VERSION : 0.1
   VAR_INPUT
      Ir_Pos_1 : Bool;   // Comando Mover Cilindro a Posición 1, activar constantemente
      Ir_Pos_2 : Bool;   // Comando Mover Cilindro a Posición 2, activar constantemente
      Conf_Pos_1 : Bool;   // Confirmación Cilindro en Posición 1
      Conf_Pos_2 : Bool;   // Confirmación Cilindro en Posición 2
      T_Conf : Time := T#10s;   // Tiempo admisible para confirmación de posición
      T_ON : Time;   // Duración accionamiento salida [0 = constantemente]
   END_VAR
   VAR_OUTPUT
      Pos_1 : Bool;   // Orden Mover Cilindro a Posición 1
      Pos_2 : Bool;   // Orden Mover Cilindro a Posición 2
      ERROR : Int;   // 0 = Sin Error, 1 = Error Programación, 2 = Error Doble Confirmación, 3 = Error Confirmación Pos_1, 4 = Error Confirmación Pos_2, 5 = Sin Confirmaciones
   END_VAR
   VAR
      IEC_Timer_0_Instance : IEC_TIMER;
      IEC_Timer_0_Instance_1 : IEC_TIMER;
      IEC_Timer_0_Instance_2 : IEC_TIMER;
      IEC_Timer_0_Instance_3 : IEC_TIMER;
      IEC_Timer_0_Instance_4 : IEC_TIMER;
   END_VAR
   VAR_TEMP
      Aux_1 : Bool;   // Auxiliar 1
      Aux_2 : Bool;   // Auxiliar 2
      Aux_ERROR : Int;   // Auxiliar ERROR
   END_VAR
BEGIN

REGION Network 1: Auxiliar 1
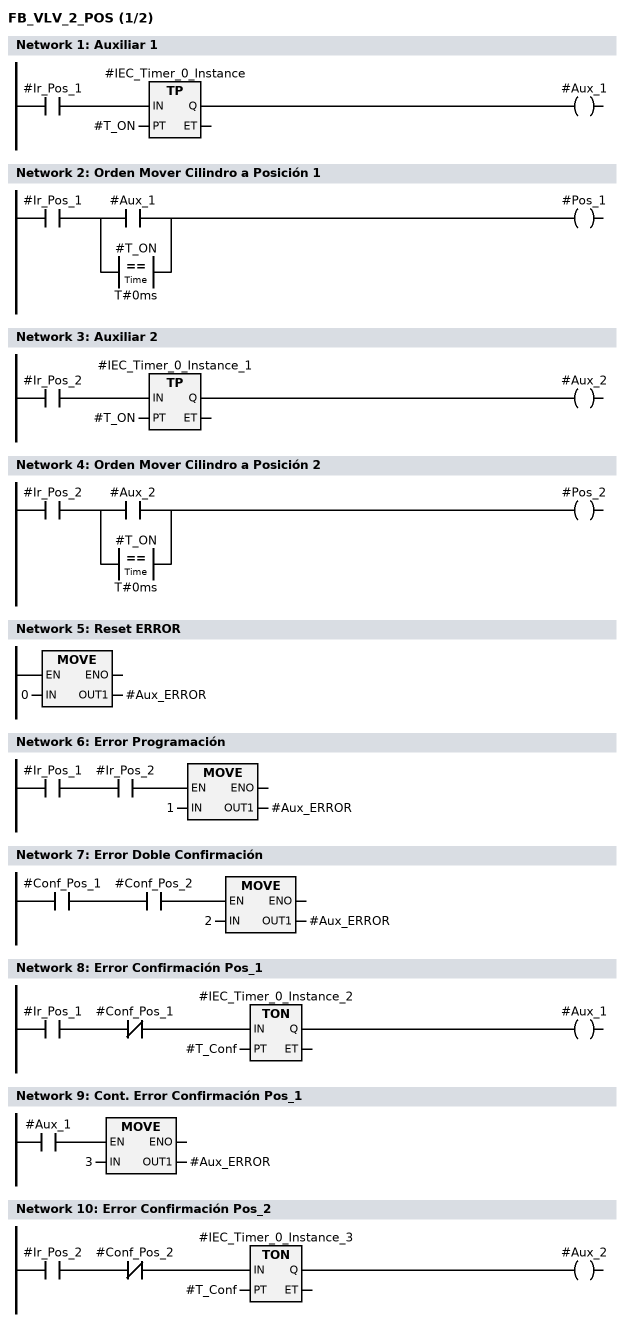
   #IEC_Timer_0_Instance.TP(IN := #Ir_Pos_1, PT := #T_ON);
   #Aux_1 := #IEC_Timer_0_Instance.Q;
END_REGION

REGION Network 2: Orden Mover Cilindro a Posición 1
   RUNG wire#powerrail
      Contact( #Ir_Pos_1 )
      wire#w1
      Contact( #Aux_1 )
      wire#w2
      Coil( #Pos_1 )
   END_RUNG
   RUNG wire#w1
      { S7_Templates := "SrcType := Time" } EQ_Contact(in1 := #T_ON, in2 := T#0ms)
   END_RUNG wire#w2
   // the same network as SCL:
   #Pos_1 := #Ir_Pos_1 AND (#Aux_1 OR (#T_ON = T#0ms));
END_REGION

REGION Network 3: Auxiliar 2
   #IEC_Timer_0_Instance_1.TP(IN := #Ir_Pos_2, PT := #T_ON);
   #Aux_2 := #IEC_Timer_0_Instance_1.Q;
END_REGION

REGION Network 4: Orden Mover Cilindro a Posición 2
   RUNG wire#powerrail
      Contact( #Ir_Pos_2 )
      wire#w1
      Contact( #Aux_2 )
      wire#w2
      Coil( #Pos_2 )
   END_RUNG
   RUNG wire#w1
      { S7_Templates := "SrcType := Time" } EQ_Contact(in1 := #T_ON, in2 := T#0ms)
   END_RUNG wire#w2
   // the same network as SCL:
   #Pos_2 := #Ir_Pos_2 AND (#Aux_2 OR (#T_ON = T#0ms));
END_REGION

REGION Network 5: Reset ERROR
   RUNG wire#powerrail
      { S7_GenerateENO := "TRUE" } Move(in := 0, out1 => #Aux_ERROR)
   END_RUNG
   // the same network as SCL:
   #Aux_ERROR := 0;
END_REGION

REGION Network 6: Error Programación
   RUNG wire#powerrail
      Contact( #Ir_Pos_1 )
      Contact( #Ir_Pos_2 )
      { S7_GenerateENO := "TRUE" } Move(in := 1, out1 => #Aux_ERROR)
   END_RUNG
   // the same network as SCL:
   IF #Ir_Pos_1 AND #Ir_Pos_2 THEN #Aux_ERROR := 1; END_IF;
END_REGION

REGION Network 7: Error Doble Confirmación
   RUNG wire#powerrail
      Contact( #Conf_Pos_1 )
      Contact( #Conf_Pos_2 )
      { S7_GenerateENO := "TRUE" } Move(in := 2, out1 => #Aux_ERROR)
   END_RUNG
   // the same network as SCL:
   IF #Conf_Pos_1 AND #Conf_Pos_2 THEN #Aux_ERROR := 2; END_IF;
END_REGION

REGION Network 8: Error Confirmación Pos_1
   #IEC_Timer_0_Instance_2.TON(IN := #Ir_Pos_1 AND NOT #Conf_Pos_1, PT := #T_Conf);
   #Aux_1 := #IEC_Timer_0_Instance_2.Q;
END_REGION

REGION Network 9: Cont. Error Confirmación Pos_1
   RUNG wire#powerrail
      Contact( #Aux_1 )
      { S7_GenerateENO := "TRUE" } Move(in := 3, out1 => #Aux_ERROR)
   END_RUNG
   // the same network as SCL:
   IF #Aux_1 THEN #Aux_ERROR := 3; END_IF;
END_REGION

REGION Network 10: Error Confirmación Pos_2
   #IEC_Timer_0_Instance_3.TON(IN := #Ir_Pos_2 AND NOT #Conf_Pos_2, PT := #T_Conf);
   #Aux_2 := #IEC_Timer_0_Instance_3.Q;
END_REGION

REGION Network 11: Cont. Error Confirmación Pos_2
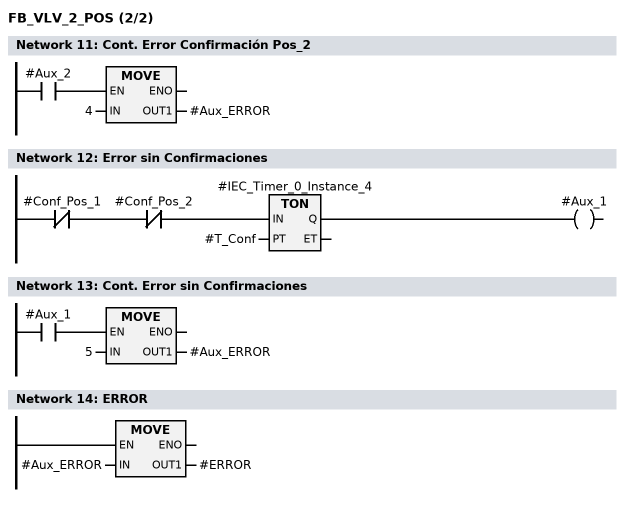
   RUNG wire#powerrail
      Contact( #Aux_2 )
      { S7_GenerateENO := "TRUE" } Move(in := 4, out1 => #Aux_ERROR)
   END_RUNG
   // the same network as SCL:
   IF #Aux_2 THEN #Aux_ERROR := 4; END_IF;
END_REGION

REGION Network 12: Error sin Confirmaciones
   #IEC_Timer_0_Instance_4.TON(IN := NOT #Conf_Pos_1 AND NOT #Conf_Pos_2, PT := #T_Conf);
   #Aux_1 := #IEC_Timer_0_Instance_4.Q;
END_REGION

REGION Network 13: Cont. Error sin Confirmaciones
   RUNG wire#powerrail
      Contact( #Aux_1 )
      { S7_GenerateENO := "TRUE" } Move(in := 5, out1 => #Aux_ERROR)
   END_RUNG
   // the same network as SCL:
   IF #Aux_1 THEN #Aux_ERROR := 5; END_IF;
END_REGION

REGION Network 14: ERROR
   RUNG wire#powerrail
      { S7_GenerateENO := "TRUE" } Move(in := #Aux_ERROR, out1 => #ERROR)
   END_RUNG
   // the same network as SCL:
   #ERROR := #Aux_ERROR;
END_REGION
END_FUNCTION_BLOCK

FUNCTION "MAQ_EST_32" : Void   // FC7, SCL
TITLE = Máquina de Estados 32
{ S7_Optimized_Access := 'TRUE' }
AUTHOR : FRD
FAMILY : MTA
NAME : MaqEst32
VERSION : 1.0
// KNOW_HOW_PROTECT  Máquina de estados de hasta 32 estados.
   VAR_INPUT
      Concatenadoras : DWord;   // Próximo estado de transición normal
      Prioritarias : DWord;   // Próximo estado de transición forzada
   END_VAR
   VAR_OUTPUT
      Error_Concatenadoras : Bool;   // Error en la programación de las Concatenadoras
      Error_Prioritarias : Bool;   // Error en la programación de las Prioritarias
   END_VAR
   VAR_IN_OUT
      Estado : DWord;   // Estado actual
   END_VAR
   VAR_TEMP
      Concat_Int : Int;   // Auxiliar INT para verificar las Concatenadoras
      Priorit_Int : Int;   // Auxiliar INT para verificar las Prioritarias
      Concat_Dword : DWord;   // Auxiliar DWORD para verificar las Concatenadoras
      Priorit_Dword : DWord;   // Auxiliar DWORD para verificar las Prioritarias
      Activar_Concat : Bool;   // Bit que indica Concatenadoras correctas
      Activar_Priorit : Bool;   // Bit que indica Prioritarias correctas
      Falla_Concat : Bool;   // Bit que indica falla en Concatenadoras
      Falla_Priorit : Bool;   // Bit que indica falla en Prioritarias
   END_VAR
BEGIN
   #Falla_Concat := 0;
   #Activar_Concat := 0;
   #Falla_Priorit := 0;
   #Activar_Priorit := 0; 
   #Error_Concatenadoras := 0;
   #Error_Prioritarias := 0;

   IF #Concatenadoras <> 0 THEN     //Evaluar Concatenadoras si son distintas de "0"

    #Concat_Int := ENCO(IN := #Concatenadoras );  //Convierte posición_DWORD en INT (0 a 31), lee el LSb

    #Concat_Dword := DECO(IN := INT_TO_UINT(#Concat_Int));//Convierte INT en posición_DWORD (1 a 32)

    IF #Concatenadoras = #Concat_Dword THEN  //Si son iguales, había sólo un bit en "1"

     #Activar_Concat := 1;    //Concatenadora correcta

    ELSE

     #Falla_Concat := 1;    //Falla en Concatenadora

    END_IF;

   END_IF;

   IF #Prioritarias <> 0 THEN     //Evaluar Prioritarias si son distintas de "0"

    #Priorit_Int := ENCO(IN := #Prioritarias);  //Convierte posición_DWORD en INT (0 a 31), lee el LSb

    #Priorit_Dword := DECO(IN := INT_TO_UINT(#Priorit_Int));//Convierte INT en posición_DWORD (1 a 32)

    IF #Prioritarias = #Priorit_Dword THEN  //Si son iguales, había sólo un bit en "1"

     #Activar_Priorit := 1;   //Prioritaria correcta

    ELSE

     #Falla_Priorit := 1;    //Falla en Prioritaria

    END_IF;

   END_IF;

   IF NOT(#Falla_Priorit OR #Falla_Concat) THEN  //Si no hay falla de Prioritaria ni de Concatenadora

    IF #Activar_Priorit THEN    //Si hay que asignar Prioritarias

     #Estado := #Prioritarias;

    ELSE

     IF #Activar_Concat THEN   //Si hay que asignar Concatenadoras

      #Estado := #Concatenadoras;

     END_IF;

    END_IF;

   ELSE

    IF #Falla_Concat THEN     //Si hay falla de Concatenadoras

     #Error_Concatenadoras := 1;    //Activar Error_Concatenadoras

    END_IF;

    IF #Falla_Priorit THEN    //Si hay falla de Prioritarias

     #Error_Prioritarias := 1;    //Activar Error_Prioritarias

    END_IF;

   END_IF;
END_FUNCTION

// folder: INCIDENTES

FUNCTION_BLOCK "FB_INC_GENERAL"   // FB500, LAD
TITLE = ALARMAS GENERAL
{ S7_Optimized_Access := 'FALSE' }
VERSION : 0.1
   VAR
      Alarma_On : Bool;
   END_VAR
BEGIN

REGION Network 1: Alarma 0 - Protecciones abiertas
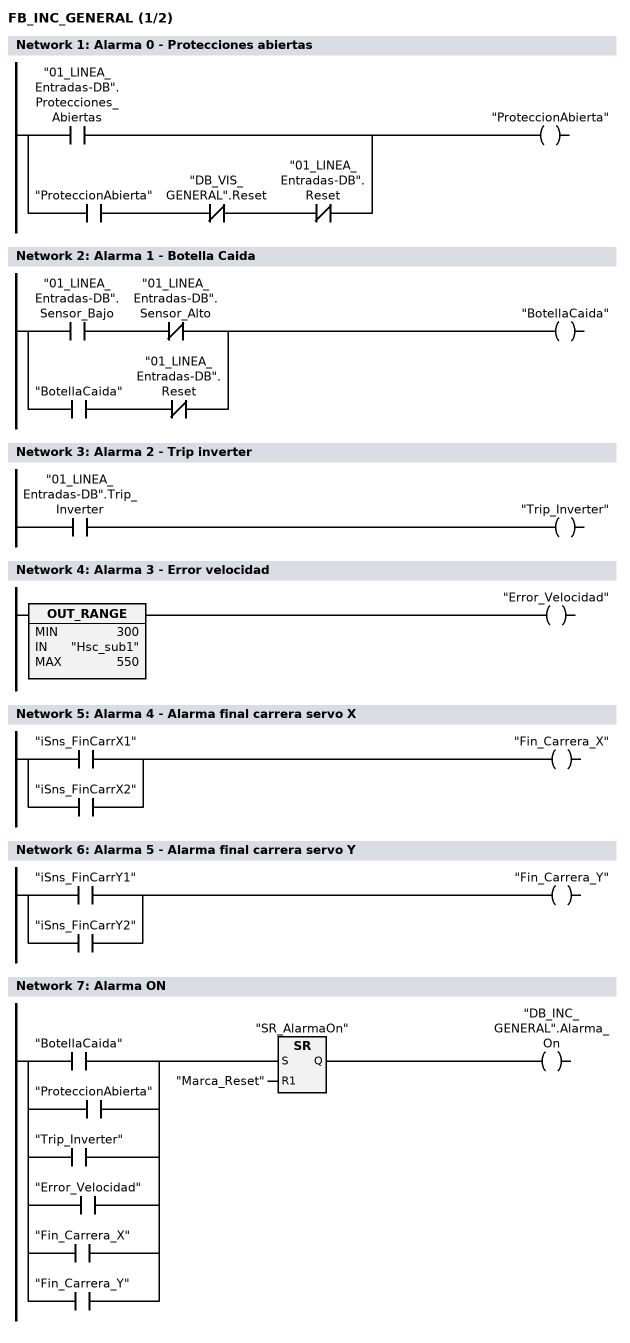
   RUNG wire#powerrail
      Contact( "01_LINEA_Entradas-DB".Protecciones_Abiertas )
      wire#w1
      Coil( "ProteccionAbierta" )
   END_RUNG
   RUNG wire#powerrail
      Contact( "ProteccionAbierta" )
      I_Contact( "DB_VIS_GENERAL".Reset )
      I_Contact( "01_LINEA_Entradas-DB".Reset )
   END_RUNG wire#w1
   // the same network as SCL:
   "ProteccionAbierta" := "01_LINEA_Entradas-DB".Protecciones_Abiertas OR ("ProteccionAbierta" AND NOT "DB_VIS_GENERAL".Reset AND NOT "01_LINEA_Entradas-DB".Reset);
END_REGION

REGION Network 2: Alarma 1 - Botella Caida
   RUNG wire#powerrail
      Contact( "01_LINEA_Entradas-DB".Sensor_Bajo )
      I_Contact( "01_LINEA_Entradas-DB".Sensor_Alto )
      wire#w1
      Coil( "BotellaCaida" )
   END_RUNG
   RUNG wire#powerrail
      Contact( "BotellaCaida" )
      I_Contact( "01_LINEA_Entradas-DB".Reset )
   END_RUNG wire#w1
   // the same network as SCL:
   "BotellaCaida" := ("01_LINEA_Entradas-DB".Sensor_Bajo AND NOT "01_LINEA_Entradas-DB".Sensor_Alto) OR ("BotellaCaida" AND NOT "01_LINEA_Entradas-DB".Reset);
END_REGION

REGION Network 3: Alarma 2 - Trip inverter
   RUNG wire#powerrail
      Contact( "01_LINEA_Entradas-DB".Trip_Inverter )
      Coil( "Trip_Inverter" )
   END_RUNG
   // the same network as SCL:
   "Trip_Inverter" := "01_LINEA_Entradas-DB".Trip_Inverter;
END_REGION

REGION Network 4: Alarma 3 - Error velocidad
   "Error_Velocidad" := ("Hsc_sub1" < 300) OR ("Hsc_sub1" > 550);
END_REGION

REGION Network 5: Alarma 4 - Alarma final carrera servo X
   RUNG wire#powerrail
      Contact( "iSns_FinCarrX1" )
      wire#w1
      Coil( "Fin_Carrera_X" )
   END_RUNG
   RUNG wire#powerrail
      Contact( "iSns_FinCarrX2" )
   END_RUNG wire#w1
   // the same network as SCL:
   "Fin_Carrera_X" := "iSns_FinCarrX1" OR "iSns_FinCarrX2";
END_REGION

REGION Network 6: Alarma 5 - Alarma final carrera servo Y
   RUNG wire#powerrail
      Contact( "iSns_FinCarrY1" )
      wire#w1
      Coil( "Fin_Carrera_Y" )
   END_RUNG
   RUNG wire#powerrail
      Contact( "iSns_FinCarrY2" )
   END_RUNG wire#w1
   // the same network as SCL:
   "Fin_Carrera_Y" := "iSns_FinCarrY1" OR "iSns_FinCarrY2";
END_REGION

REGION Network 7: Alarma ON
   RUNG wire#powerrail
      Contact( "BotellaCaida" )
      wire#w1
      S_SR(operand := "SR_AlarmaOn", r1 := "Marca_Reset")
      Coil( "DB_INC_GENERAL".Alarma_On )
   END_RUNG
   RUNG wire#powerrail
      Contact( "ProteccionAbierta" )
   END_RUNG wire#w1
   RUNG wire#powerrail
      Contact( "Trip_Inverter" )
   END_RUNG wire#w1
   RUNG wire#powerrail
      Contact( "Error_Velocidad" )
   END_RUNG wire#w1
   RUNG wire#powerrail
      Contact( "Fin_Carrera_X" )
   END_RUNG wire#w1
   RUNG wire#powerrail
      Contact( "Fin_Carrera_Y" )
   END_RUNG wire#w1
   // the same network as SCL:
   IF "BotellaCaida" OR "ProteccionAbierta" OR "Trip_Inverter" OR "Error_Velocidad" OR "Fin_Carrera_X" OR "Fin_Carrera_Y" THEN
       "SR_AlarmaOn" := TRUE;   // SR flip-flop
   END_IF;
   IF "Marca_Reset" THEN "SR_AlarmaOn" := FALSE; END_IF;
   "DB_INC_GENERAL".Alarma_On := "SR_AlarmaOn";
END_REGION

REGION Network 8: Encendido Semaforo Rojo
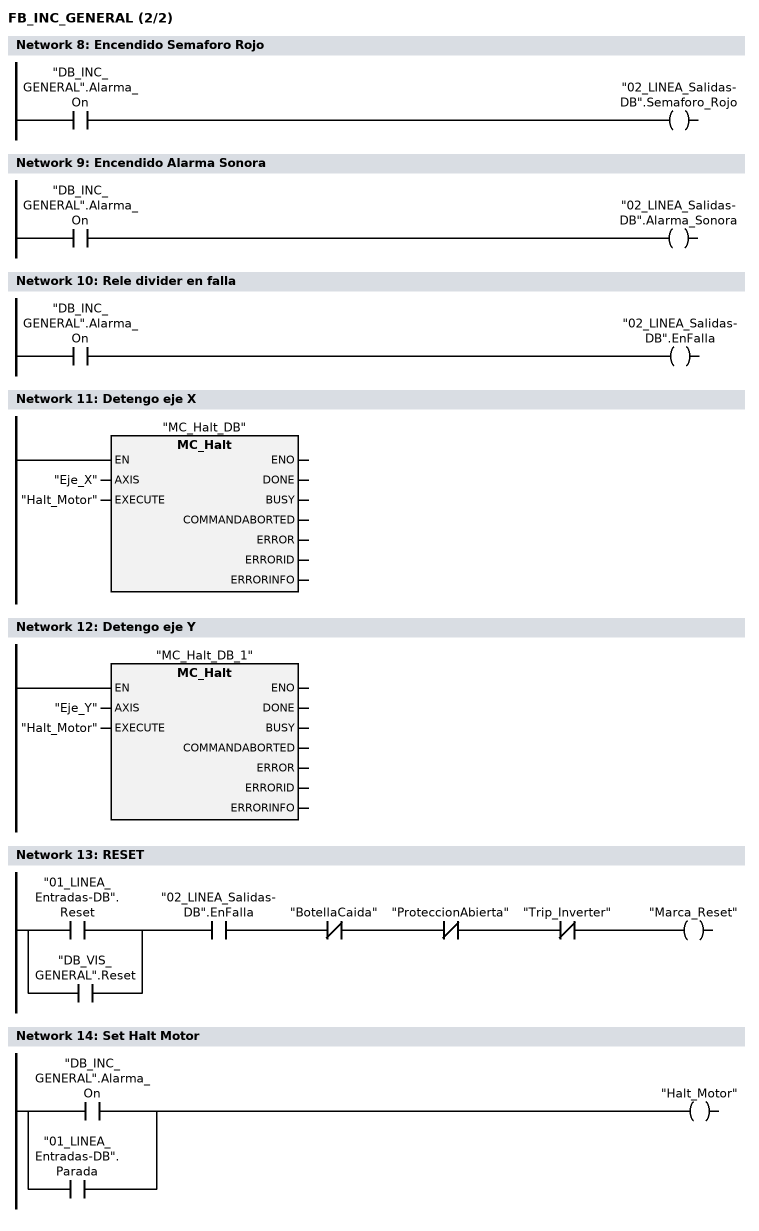
   RUNG wire#powerrail
      Contact( "DB_INC_GENERAL".Alarma_On )
      Coil( "02_LINEA_Salidas-DB".Semaforo_Rojo )
   END_RUNG
   // the same network as SCL:
   "02_LINEA_Salidas-DB".Semaforo_Rojo := "DB_INC_GENERAL".Alarma_On;
END_REGION

REGION Network 9: Encendido Alarma Sonora
   RUNG wire#powerrail
      Contact( "DB_INC_GENERAL".Alarma_On )
      Coil( "02_LINEA_Salidas-DB".Alarma_Sonora )
   END_RUNG
   // the same network as SCL:
   "02_LINEA_Salidas-DB".Alarma_Sonora := "DB_INC_GENERAL".Alarma_On;
END_REGION

REGION Network 10: Rele divider en falla
   RUNG wire#powerrail
      Contact( "DB_INC_GENERAL".Alarma_On )
      Coil( "02_LINEA_Salidas-DB".EnFalla )
   END_RUNG
   // the same network as SCL:
   "02_LINEA_Salidas-DB".EnFalla := "DB_INC_GENERAL".Alarma_On;
END_REGION

REGION Network 11: Detengo eje X
   "MC_Halt_DB"(Axis := "Eje_X", Execute := "Halt_Motor");   // MC_Halt
END_REGION

REGION Network 12: Detengo eje Y
   "MC_Halt_DB_1"(Axis := "Eje_Y", Execute := "Halt_Motor");   // MC_Halt
END_REGION

REGION Network 13: RESET
   RUNG wire#powerrail
      Contact( "01_LINEA_Entradas-DB".Reset )
      wire#w1
      Contact( "02_LINEA_Salidas-DB".EnFalla )
      I_Contact( "BotellaCaida" )
      I_Contact( "ProteccionAbierta" )
      I_Contact( "Trip_Inverter" )
      Coil( "Marca_Reset" )
   END_RUNG
   RUNG wire#powerrail
      Contact( "DB_VIS_GENERAL".Reset )
   END_RUNG wire#w1
   // the same network as SCL:
   "Marca_Reset" := ("01_LINEA_Entradas-DB".Reset OR "DB_VIS_GENERAL".Reset) AND "02_LINEA_Salidas-DB".EnFalla AND NOT "BotellaCaida" AND NOT "ProteccionAbierta" AND NOT "Trip_Inverter";
END_REGION

REGION Network 14: Set Halt Motor
   RUNG wire#powerrail
      Contact( "DB_INC_GENERAL".Alarma_On )
      wire#w1
      Coil( "Halt_Motor" )
   END_RUNG
   RUNG wire#powerrail
      Contact( "01_LINEA_Entradas-DB".Parada )
   END_RUNG wire#w1
   // the same network as SCL:
   "Halt_Motor" := "DB_INC_GENERAL".Alarma_On OR "01_LINEA_Entradas-DB".Parada;
END_REGION
END_FUNCTION_BLOCK

(* ===== HMI "HMI_RT_1" =====
system functions are stored by id; their names below are inferred from use
connection "Conexión_1": ETHERNET, SMART_S7_1200_OMS
connection "HMI_Conexión_1": ETHERNET, SMART_S7_1200_OMS

HMI tags "Tabla de variables estándar"
   "MC_Power_X" : Bool = PLC DB_VIS_GENERAL.MC_Pwr_EnX AT %DB800.DBX2.2, 1 s
   "MC_Power_Y" : Bool = PLC DB_VIS_GENERAL.MC_Pwrt_EnY AT %DB800.DBX2.3, 1 s
   "MC_JogFwd_X" : Bool = PLC DB_VIS_GENERAL.MC_JogFwd_X AT %DB800.DBX2.6, 1 s
   "MC_JogFwd_Y" : Bool = PLC DB_VIS_GENERAL.MC_JogFwd_Y AT %DB800.DBX2.7, 1 s
   "MC_JogBckWd_X" : Bool = PLC DB_VIS_GENERAL.MC_JogBwd_X AT %DB800.DBX3.0, 1 s
   "MC_JogBckWd_Y" : Bool = PLC DB_VIS_GENERAL.MC_JogBwd_Y AT %DB800.DBX3.1, 1 s
   "Falla_Divider" : Bool = PLC "02_LINEA_Salidas-DB".EnFalla AT %DB1.DBX0.0, 1 s
   "ProteccionesAbiertas" : Bool = PLC "01_LINEA_Entradas-DB".Protecciones_Abiertas AT %DB1.DBX0.0, 1 s
   "BotellaCaida" : Bool = PLC BotellaCaida AT %M100.1, 1 s
   "Marcha_Divider" : Bool = PLC "02_LINEA_Salidas-DB".EnMarcha AT %DB1.DBX0.0, 1 s
   "Trip_Inverter" : Bool = PLC Trip_Inverter AT %M100.2, 1 s
   "Cant_Bot" : Int = PLC DB_VIS_GENERAL.CantBot AT %DB800.DBW0, 1 s
   "Marcha" : Bool = PLC DB_VIS_GENERAL.Start AT %DB800.DBX3.4, 1 s
   "HomingOk" : Bool = PLC DB_VIS_GENERAL.HomingOk AT %DB800.DBX3.2, 1 s
   "Reset" : Bool = PLC DB_VIS_GENERAL.Reset AT %DB800.DBX3.3, 1 s
   "PM_MovX" : Real = PLC DB_PUESTA_MARCHA.MovXmm AT %DB1.DBX0.0, 1 s
   "PM_MovY" : Real = PLC DB_PUESTA_MARCHA.MovYmm AT %DB1.DBX0.0, 1 s
   "PM_TChFull" : Time = PLC DB_PUESTA_MARCHA.TChFull AT %DB1.DBX0.0, 1 s
   "Alarmas_1" : Word = PLC Alarmas_1 AT %MW100, 1 s
   "Alarma_ON" : Bool = PLC DB_INC_GENERAL.Alarma_On AT %DB500.DBX0.0, 1 s

discrete alarms
   1: 'Alarma 0 - Protecciones abiertas', class Errors, trigger "Alarmas_1" bit 8
   2: 'Alarma 1 - Botella caida', class Errors, trigger "Alarmas_1" bit 9
   3: 'Alarma 2 - Trip Inverter', class Errors, trigger "Alarmas_1" bit 10
   4: 'Alarma 3 - Error de velocidad', class Errors, trigger "Alarmas_1" bit 11
   5: 'Alarma 4 - Final de carrera X', class Errors, trigger "Alarmas_1" bit 12
   6: 'Alarma 5 - Final de carrera Y', class Errors, trigger "Alarmas_1" bit 13

text list "Cant_Bot": 0 '0'; 2 '2'; 4 '4'; 6 '6'; 8 '8'; 10 '10'; 12 '12'; 14 '14'; 16 '16'; 18 '18'; 20 '20'

text list "DesplazamientoX": 0 '0'; 60 '60'; 20 '20'; 40 '40'

screen "02 - Estado" 800x480, template "Plantilla_1"
   Button "Botón_2" at 162,433 size 160x46; TextOff 'Fallas'
      on Click: ActivateScreen("03 - Registro alarmas", 0)
   TextField "Campo de texto_13" at 340,308 size 197x34; Text 'Divider en falla'
   GraphicIOField "PlotLight_Round_R_2" at 222,278 size 108x108; PictureOff "PilotLight_Round_R_Off_256c"; PictureOn "PilotLight_Round_R_On_256c"
      ProcessValue <- "Falla_Divider"
   GraphicIOField "PlotLight_Round_G_16" at 223,153 size 108x108; PictureOff "PilotLight_Round_G_Off_256c"; PictureOn "PilotLight_Round_G_On_256c"
      ProcessValue <- "Marcha_Divider"
   TextField "Campo de texto_14" at 340,187 size 235x34; Text 'Divider en marcha'
   Button "Botón_3" at 14,210 size 144x51; TextOff 'START'
      on Click: SetBit("Marcha")
   SymbolicIOField "Campo ES simbólico_1" at 222,81 size 104x49; TextOn '1'; TextOff '0'; TextList "Cant_Bot"
      ProcessValue <- "Cant_Bot"
   TextField "Campo de texto_2" at 340,87 size 385x34; Text 'Cantidad de botellas por carril'
   TextField "Campo de texto_1" at 10,406 size 148x17; Text 'Solo con Divider detenido'
   Button "Botón_4" at 640,431 size 159x48; TextOff 'Protegido'; Authorization "Administración de usuarios"
      on Click: ActivateScreen("04 - Puesta en marcha", 0)
   Button "Botón_1" at 1,433 size 161x47; TextOff 'Homing'
      on Click: ActivateScreen("01 - Pantalla_Inicializacion", 0)
      Visibility <- "Marcha"
   Button "Botón_5" at 2,433 size 161x47; TextOff 'Homing'
      Visibility <- "Marcha"

screen "01 - Pantalla_Inicializacion" 800x480, template "Plantilla_1"
   Button "Botón_1" at 321,432 size 161x47; TextOff 'HOMING OK'
      on Click: ActivateScreen("02 - Estado", 0); SetBit("HomingOk"); ResetBit("Reset")
   TextField "Campo de texto_1" at 49,36 size 704x94; Text '1. HABILITE AMBOS EJES 2. POSICIONE DIVIDER EN CARRIL 1 CON PULSADORES 3. PRESIONE HOMING OK UNA VEZ FINALIZADO'
   Button "FB_ArrowDown_Round" at 144,309 size 74x74; TextOff 'Text'; PictureOff "FB_ArrowDown_Round_Released_256c"; PictureOn "FB_ArrowDown_Round_Pressed_256c"
      on Release: ResetBit("MC_JogFwd_X")
      on Press: SetBit("MC_JogFwd_X")
   Button "FB_ArrowUp_Round" at 250,309 size 74x74; TextOff 'Text'; PictureOff "FB_ArrowUp_Round_Released_256c"; PictureOn "FB_ArrowUp_Round_Pressed_256c"
      on Release: ResetBit("MC_JogBckWd_X")
      on Press: SetBit("MC_JogBckWd_X")
   Button "FB_ArrowLeft_Round" at 488,308 size 74x74; TextOff 'Text'; PictureOff "FB_ArrowLeft_Round_Released_256c"; PictureOn "FB_ArrowLeft_Round_Pressed_256c"
      on Press: SetBit("MC_JogFwd_Y")
      on Release: ResetBit("MC_JogFwd_Y")
   Button "FB_ArrowRight_Round" at 594,309 size 74x74; TextOff 'Text'; PictureOff "FB_ArrowRight_Round_Released_256c"; PictureOn "FB_ArrowRight_Round_Pressed_256c"
      on Press: SetBit("MC_JogBckWd_Y")
      on Release: ResetBit("MC_JogBckWd_Y")
   Button "FB_Check_Round" at 199,199 size 74x74; TextOff 'Text'; PictureOn "FB_Check_Round_Pressed_256c"; PictureOff "FB_Check_Round_Released_256c"
      on Click: InvertBit("MC_Power_X")
      Appearance <- "MC_Power_X"
   Button "FB_Check_Round_1" at 544,199 size 74x74; TextOff 'Text'; PictureOff "FB_Check_Round_Released_256c"; PictureOn "FB_Check_Round_Pressed_256c"
      on Click: InvertBit("MC_Power_Y")
      Appearance <- "MC_Power_Y"
   TextField "Campo de texto_3" at 174,154 size 123x23; Text 'Habilitar eje X'
   TextField "Campo de texto_2" at 519,154 size 123x23; Text 'Habilitar eje Y'
   TextField "Campo de texto_4" at 372,177 size 16x23; Text 'Text'
   Button "Botón_2" at 162,433 size 160x46; TextOff 'Fallas'
      on Click: ActivateScreen("03 - Registro alarmas", 0)
   Button "Botón_4" at 640,431 size 159x48; TextOff 'Protegido'; Authorization "Administración de usuarios"
      on Click: ActivateScreen("04 - Puesta en marcha", 0)
   Button "Botón_3" at 2,433 size 160x47; TextOff 'Estado'
      on Click: ActivateScreen("02 - Estado", 0)

screen "03 - Registro alarmas" 800x480, template "Plantilla_1"
   Button "Botón_1" at 161,431 size 160x47; TextOff 'Estado'
      on Click: ActivateScreen("02 - Estado", 0)
   TextField "Campo de texto_5" at 286,300 size 16x23; Text 'Text'
   Button "Botón_3" at 321,431 size 161x48; TextOff 'Reset'
      on Click: SetBit("Reset"); ResetBit("HomingOk"); ResetBit("Marcha")
      Appearance <- "Alarma_ON"
   Button "Botón_4" at 640,431 size 159x48; TextOff 'Protegido'; Authorization "Administración de usuarios"
      on Click: ActivateScreen("04 - Puesta en marcha", 0)
   AlarmView "Visor de avisos_1" at 0,28 size 799x404
   Button "Botón_2" at 0,432 size 161x47; TextOff 'Homing'
      on Click: ActivateScreen("01 - Pantalla_Inicializacion", 0)
      Visibility <- "Marcha"
   Button "Botón_5" at 1,432 size 161x47; TextOff 'Homing'
      Visibility <- "Marcha"

screen "04 - Puesta en marcha" 800x480, template "Plantilla_1"
   IOField "Campo ES_1" at 66,114 size 101x53; FormatPattern s999999999.999
      ProcessValue <- "PM_MovX"
   IOField "Campo ES_2" at 66,186 size 101x53; FormatPattern s999999999.999
      ProcessValue <- "PM_MovY"
   IOField "Campo ES_3" at 66,258 size 101x53; FormatPattern s9999999999
      ProcessValue <- "PM_TChFull"
   TextField "Campo de texto_1" at 193,129 size 141x23; Text 'Movimiento en X'
   TextField "Campo de texto_2" at 193,197 size 141x23; Text 'Movimiento en Y'
   TextField "Campo de texto_3" at 193,265 size 286x23; Text 'Tiempo de espera para canal lleno'
   Button "Botón_1" at 199,431 size 99x48; TextOff 'Est'
      on Click: ActivateScreen("02 - Estado", 0)

Template "Plantilla_1" 800x480
   DateTimeField "Plantilla_Campo de fecha y hora_1" at 596,2 size 197x24
   GraphicView "Plantilla_Visor de gráficos_1" at 9,2 size 76x24; Picture "eProC Logo Paneles Parte B"
*)